(* Logix 5000 project; controller FV vendor 1 type 14 code 217 rev 31.11; software revision 31.00; part 24 of 63 *)
(* tags used below, declared in another part *)
   CheckTimeMask : INT;
   Delphi_Does_Eng_Func : BOOL;
   FR_FV30_AV01 : PlantItem;   // FV30_AV01
   FR_FV30_AV04 : PlantItem;   // FV30_AV04
   FR_FV30_AV05 : PlantItem;   // FV30_AV05
   FR_FV30_AV06 : PlantItem;   // FV30_AV06
   FR_FV30_AV07 : PlantItem;   // FV30_AV07
   FR_FV31_AV01 : PlantItem;   // FV31_AV01
   FR_N255 : INT[265];   // CHECKWORDS
   FR_VB4_AV17 : PlantItem;   // VB4_AV17
   FR_VB4_AV18 : PlantItem;   // VB4_AV18
   FR_VB4_AV19 : PlantItem;   // VB4_AV19
   FR_VB4_AV20 : PlantItem;   // VB4_AV20
   FR_VB4_AV21 : PlantItem;   // VB4_AV21
   FR_VB4_AV22 : PlantItem;   // VB4_AV22
   FR_VB4_AV23 : PlantItem;   // VB4_AV23
   TempChecktime : DINT;
(* FR_Common, continued *)

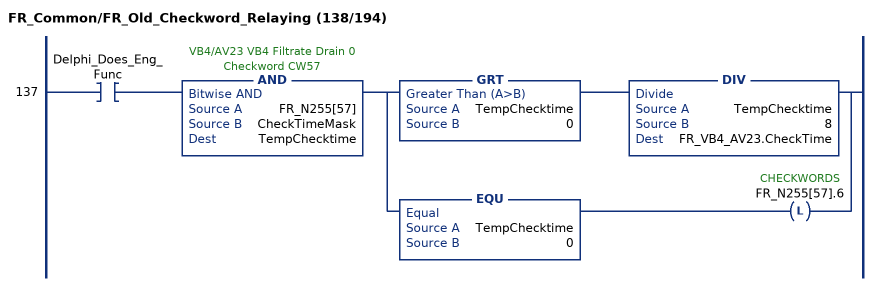
   [picture p442: FR_Common/FR_Old_Checkword_Relaying rungs 137-137]
   137: XIC(Delphi_Does_Eng_Func)AND(FR_N255[57],CheckTimeMask,TempChecktime)[GRT(TempChecktime,0) DIV(TempChecktime,8,FR_VB4_AV23.CheckTime) ,EQU(TempChecktime,0) OTL(FR_N255[57].6) ];
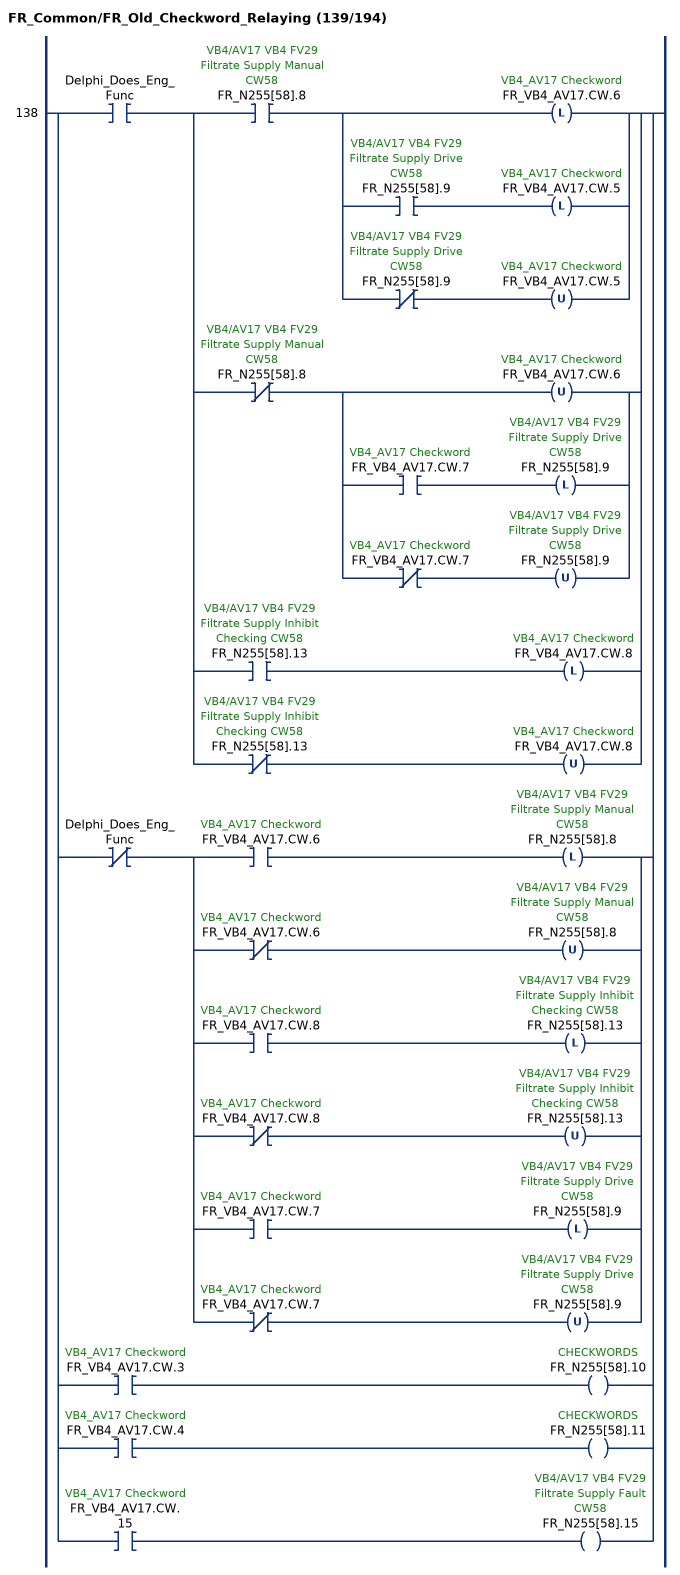
   138: [XIC(Delphi_Does_Eng_Func) [[XIC(FR_N255[58].8) [OTL(FR_VB4_AV17.CW.6) ,XIC(FR_N255[58].9) OTL(FR_VB4_AV17.CW.5) ,XIO(FR_N255[58].9) OTU(FR_VB4_AV17.CW.5) ] ,XIO(FR_N255[58].8) [OTU(FR_VB4_AV17.CW.6) ,[XIC(FR_VB4_AV17.CW.7) OTL(FR_N255[58].9) ,XIO(FR_VB4_AV17.CW.7) OTU(FR_N255[58].9) ] ] ] ,[XIC(FR_N255[58].13) OTL(FR_VB4_AV17.CW.8) ,XIO(FR_N255[58].13) OTU(FR_VB4_AV17.CW.8) ] ] ,XIO(Delphi_Does_Eng_Func) [[XIC(FR_VB4_AV17.CW.6) OTL(FR_N255[58].8) ,XIO(FR_VB4_AV17.CW.6) OTU(FR_N255[58].8) ] ,[XIC(FR_VB4_AV17.CW.8) OTL(FR_N255[58].13) ,XIO(FR_VB4_AV17.CW.8) OTU(FR_N255[58].13) ] ,[XIC(FR_VB4_AV17.CW.7) OTL(FR_N255[58].9) ,XIO(FR_VB4_AV17.CW.7) OTU(FR_N255[58].9) ] ] ,XIC(FR_VB4_AV17.CW.3) OTE(FR_N255[58].10) ,XIC(FR_VB4_AV17.CW.4) OTE(FR_N255[58].11) ,XIC(FR_VB4_AV17.CW.15) OTE(FR_N255[58].15) ];
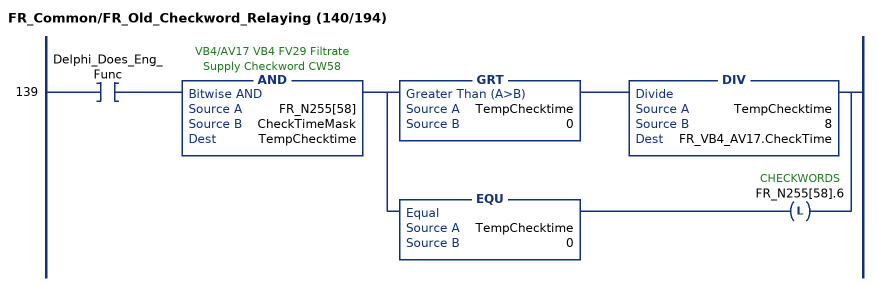
   139: XIC(Delphi_Does_Eng_Func)AND(FR_N255[58],CheckTimeMask,TempChecktime)[GRT(TempChecktime,0) DIV(TempChecktime,8,FR_VB4_AV17.CheckTime) ,EQU(TempChecktime,0) OTL(FR_N255[58].6) ];
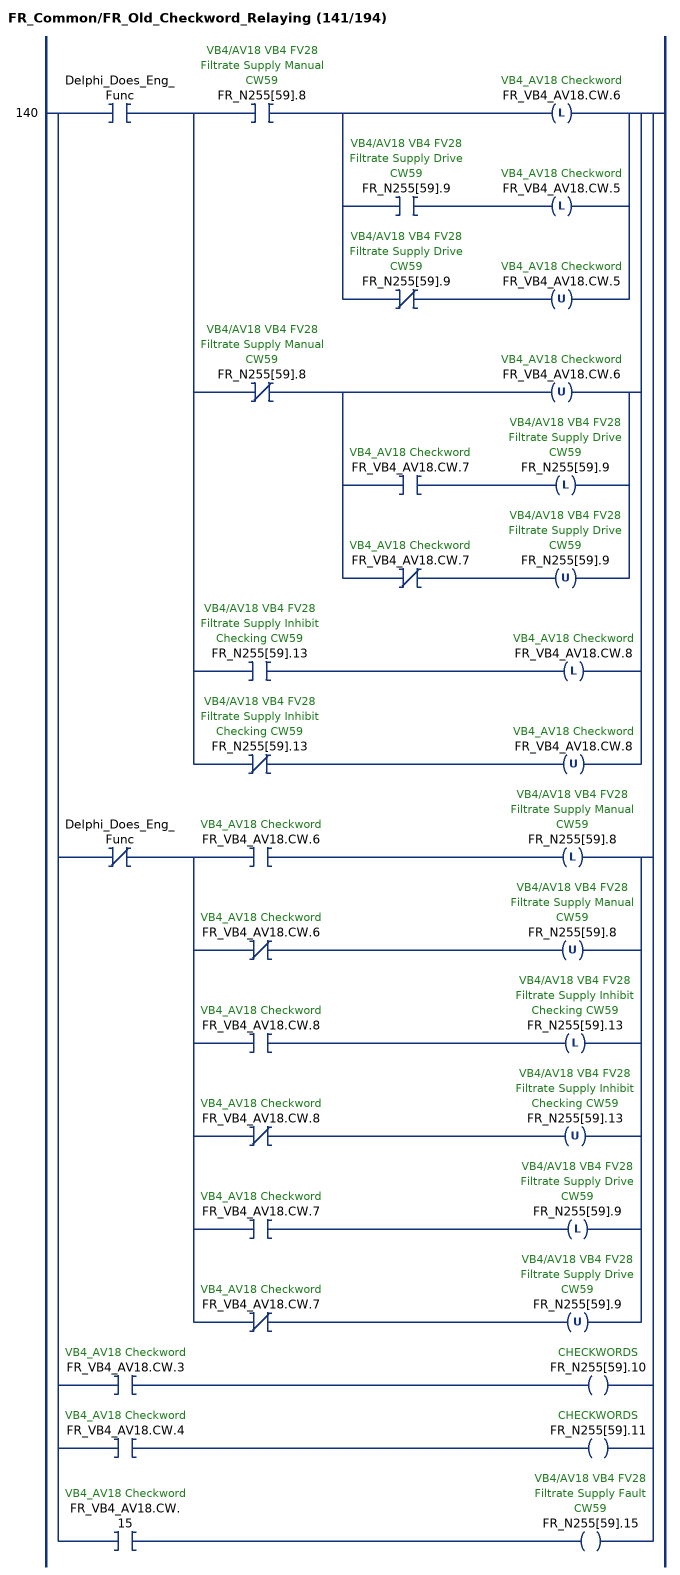
   140: [XIC(Delphi_Does_Eng_Func) [[XIC(FR_N255[59].8) [OTL(FR_VB4_AV18.CW.6) ,XIC(FR_N255[59].9) OTL(FR_VB4_AV18.CW.5) ,XIO(FR_N255[59].9) OTU(FR_VB4_AV18.CW.5) ] ,XIO(FR_N255[59].8) [OTU(FR_VB4_AV18.CW.6) ,[XIC(FR_VB4_AV18.CW.7) OTL(FR_N255[59].9) ,XIO(FR_VB4_AV18.CW.7) OTU(FR_N255[59].9) ] ] ] ,[XIC(FR_N255[59].13) OTL(FR_VB4_AV18.CW.8) ,XIO(FR_N255[59].13) OTU(FR_VB4_AV18.CW.8) ] ] ,XIO(Delphi_Does_Eng_Func) [[XIC(FR_VB4_AV18.CW.6) OTL(FR_N255[59].8) ,XIO(FR_VB4_AV18.CW.6) OTU(FR_N255[59].8) ] ,[XIC(FR_VB4_AV18.CW.8) OTL(FR_N255[59].13) ,XIO(FR_VB4_AV18.CW.8) OTU(FR_N255[59].13) ] ,[XIC(FR_VB4_AV18.CW.7) OTL(FR_N255[59].9) ,XIO(FR_VB4_AV18.CW.7) OTU(FR_N255[59].9) ] ] ,XIC(FR_VB4_AV18.CW.3) OTE(FR_N255[59].10) ,XIC(FR_VB4_AV18.CW.4) OTE(FR_N255[59].11) ,XIC(FR_VB4_AV18.CW.15) OTE(FR_N255[59].15) ];
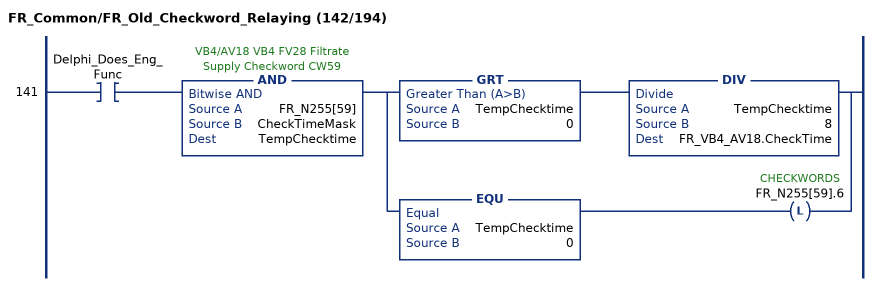
   141: XIC(Delphi_Does_Eng_Func)AND(FR_N255[59],CheckTimeMask,TempChecktime)[GRT(TempChecktime,0) DIV(TempChecktime,8,FR_VB4_AV18.CheckTime) ,EQU(TempChecktime,0) OTL(FR_N255[59].6) ];
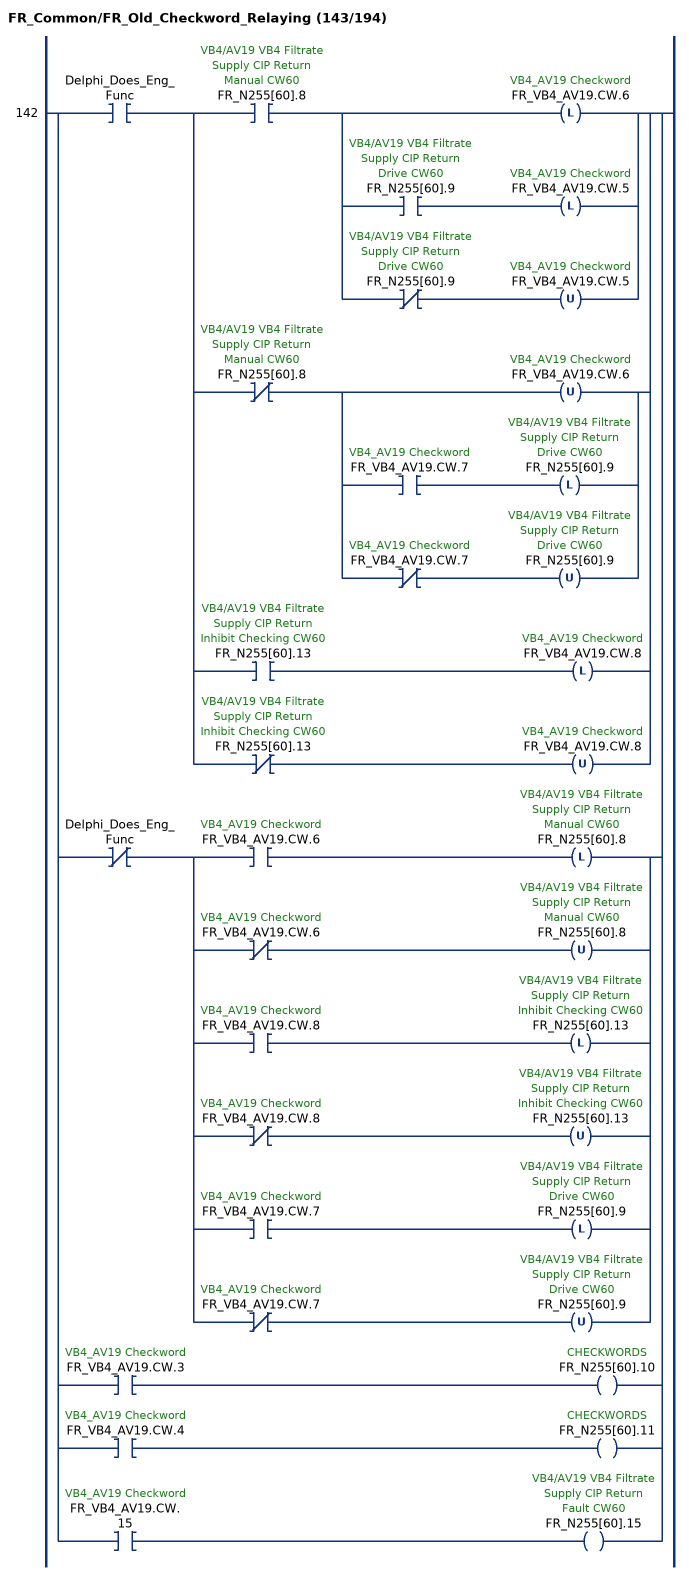
   142: [XIC(Delphi_Does_Eng_Func) [[XIC(FR_N255[60].8) [OTL(FR_VB4_AV19.CW.6) ,XIC(FR_N255[60].9) OTL(FR_VB4_AV19.CW.5) ,XIO(FR_N255[60].9) OTU(FR_VB4_AV19.CW.5) ] ,XIO(FR_N255[60].8) [OTU(FR_VB4_AV19.CW.6) ,[XIC(FR_VB4_AV19.CW.7) OTL(FR_N255[60].9) ,XIO(FR_VB4_AV19.CW.7) OTU(FR_N255[60].9) ] ] ] ,[XIC(FR_N255[60].13) OTL(FR_VB4_AV19.CW.8) ,XIO(FR_N255[60].13) OTU(FR_VB4_AV19.CW.8) ] ] ,XIO(Delphi_Does_Eng_Func) [[XIC(FR_VB4_AV19.CW.6) OTL(FR_N255[60].8) ,XIO(FR_VB4_AV19.CW.6) OTU(FR_N255[60].8) ] ,[XIC(FR_VB4_AV19.CW.8) OTL(FR_N255[60].13) ,XIO(FR_VB4_AV19.CW.8) OTU(FR_N255[60].13) ] ,[XIC(FR_VB4_AV19.CW.7) OTL(FR_N255[60].9) ,XIO(FR_VB4_AV19.CW.7) OTU(FR_N255[60].9) ] ] ,XIC(FR_VB4_AV19.CW.3) OTE(FR_N255[60].10) ,XIC(FR_VB4_AV19.CW.4) OTE(FR_N255[60].11) ,XIC(FR_VB4_AV19.CW.15) OTE(FR_N255[60].15) ];
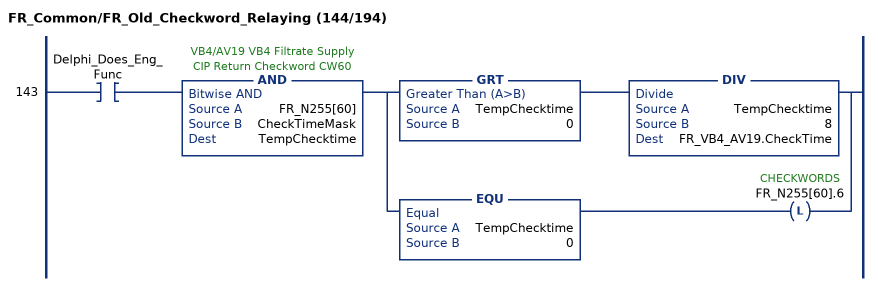
   143: XIC(Delphi_Does_Eng_Func)AND(FR_N255[60],CheckTimeMask,TempChecktime)[GRT(TempChecktime,0) DIV(TempChecktime,8,FR_VB4_AV19.CheckTime) ,EQU(TempChecktime,0) OTL(FR_N255[60].6) ];
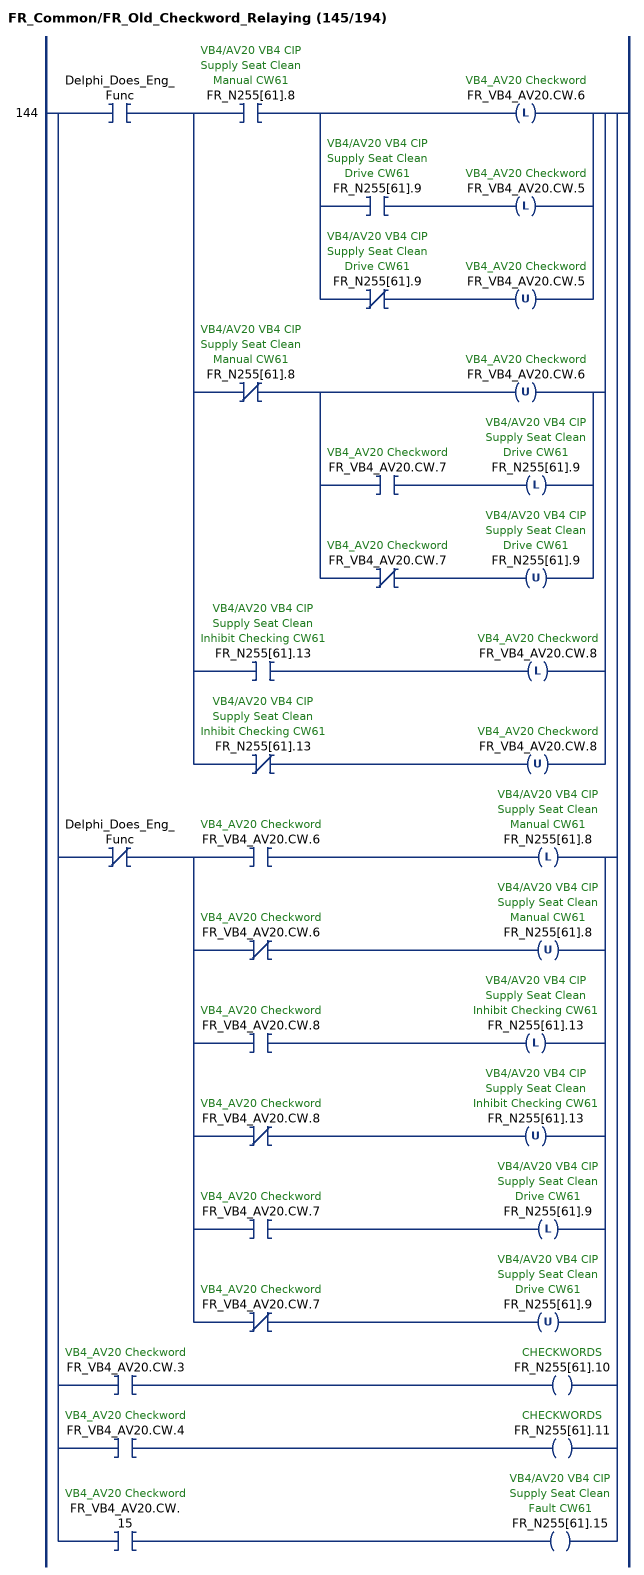
   144: [XIC(Delphi_Does_Eng_Func) [[XIC(FR_N255[61].8) [OTL(FR_VB4_AV20.CW.6) ,XIC(FR_N255[61].9) OTL(FR_VB4_AV20.CW.5) ,XIO(FR_N255[61].9) OTU(FR_VB4_AV20.CW.5) ] ,XIO(FR_N255[61].8) [OTU(FR_VB4_AV20.CW.6) ,[XIC(FR_VB4_AV20.CW.7) OTL(FR_N255[61].9) ,XIO(FR_VB4_AV20.CW.7) OTU(FR_N255[61].9) ] ] ] ,[XIC(FR_N255[61].13) OTL(FR_VB4_AV20.CW.8) ,XIO(FR_N255[61].13) OTU(FR_VB4_AV20.CW.8) ] ] ,XIO(Delphi_Does_Eng_Func) [[XIC(FR_VB4_AV20.CW.6) OTL(FR_N255[61].8) ,XIO(FR_VB4_AV20.CW.6) OTU(FR_N255[61].8) ] ,[XIC(FR_VB4_AV20.CW.8) OTL(FR_N255[61].13) ,XIO(FR_VB4_AV20.CW.8) OTU(FR_N255[61].13) ] ,[XIC(FR_VB4_AV20.CW.7) OTL(FR_N255[61].9) ,XIO(FR_VB4_AV20.CW.7) OTU(FR_N255[61].9) ] ] ,XIC(FR_VB4_AV20.CW.3) OTE(FR_N255[61].10) ,XIC(FR_VB4_AV20.CW.4) OTE(FR_N255[61].11) ,XIC(FR_VB4_AV20.CW.15) OTE(FR_N255[61].15) ];
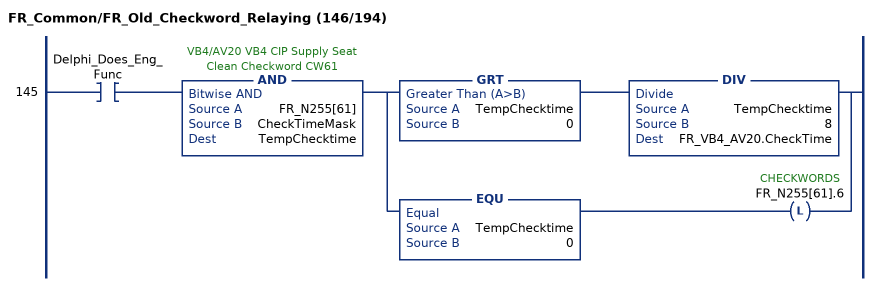
   145: XIC(Delphi_Does_Eng_Func)AND(FR_N255[61],CheckTimeMask,TempChecktime)[GRT(TempChecktime,0) DIV(TempChecktime,8,FR_VB4_AV20.CheckTime) ,EQU(TempChecktime,0) OTL(FR_N255[61].6) ];
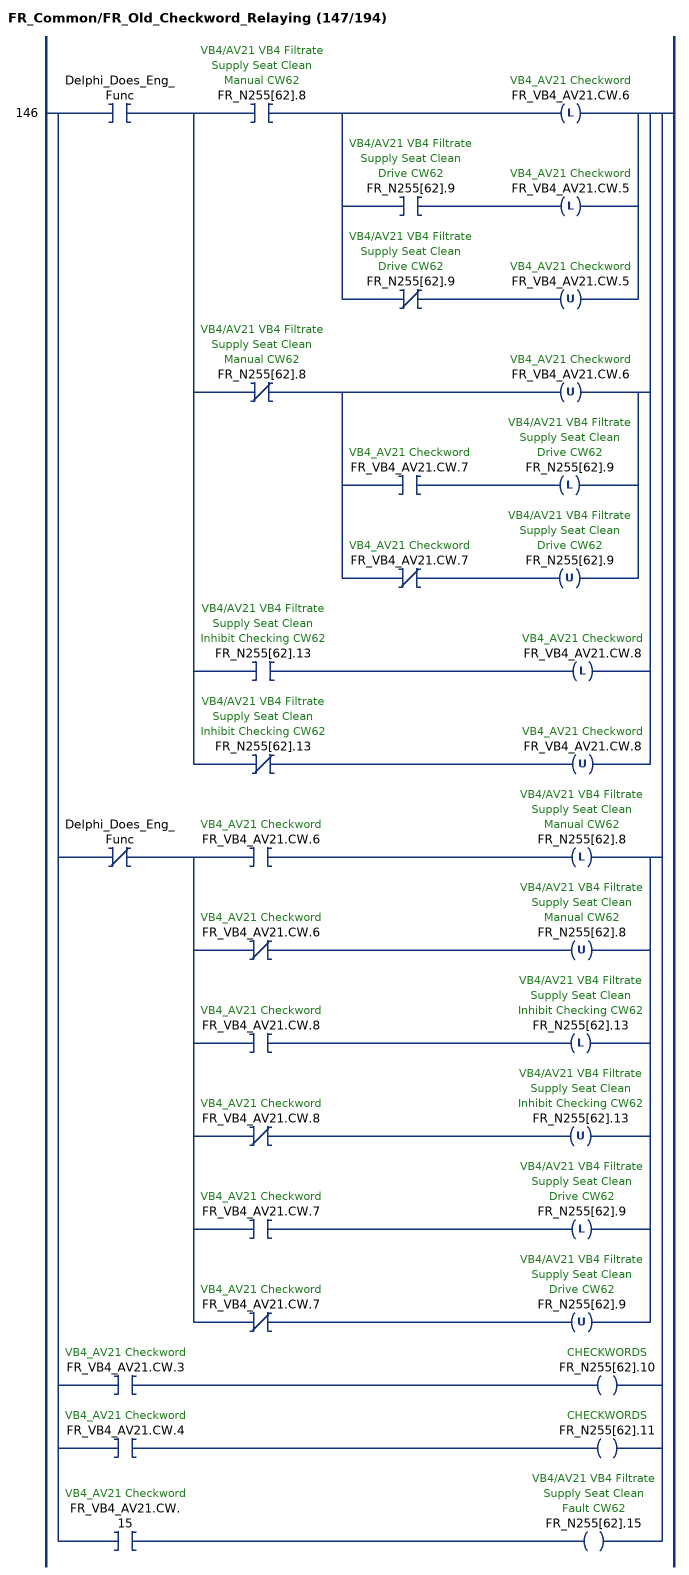
   146: [XIC(Delphi_Does_Eng_Func) [[XIC(FR_N255[62].8) [OTL(FR_VB4_AV21.CW.6) ,XIC(FR_N255[62].9) OTL(FR_VB4_AV21.CW.5) ,XIO(FR_N255[62].9) OTU(FR_VB4_AV21.CW.5) ] ,XIO(FR_N255[62].8) [OTU(FR_VB4_AV21.CW.6) ,[XIC(FR_VB4_AV21.CW.7) OTL(FR_N255[62].9) ,XIO(FR_VB4_AV21.CW.7) OTU(FR_N255[62].9) ] ] ] ,[XIC(FR_N255[62].13) OTL(FR_VB4_AV21.CW.8) ,XIO(FR_N255[62].13) OTU(FR_VB4_AV21.CW.8) ] ] ,XIO(Delphi_Does_Eng_Func) [[XIC(FR_VB4_AV21.CW.6) OTL(FR_N255[62].8) ,XIO(FR_VB4_AV21.CW.6) OTU(FR_N255[62].8) ] ,[XIC(FR_VB4_AV21.CW.8) OTL(FR_N255[62].13) ,XIO(FR_VB4_AV21.CW.8) OTU(FR_N255[62].13) ] ,[XIC(FR_VB4_AV21.CW.7) OTL(FR_N255[62].9) ,XIO(FR_VB4_AV21.CW.7) OTU(FR_N255[62].9) ] ] ,XIC(FR_VB4_AV21.CW.3) OTE(FR_N255[62].10) ,XIC(FR_VB4_AV21.CW.4) OTE(FR_N255[62].11) ,XIC(FR_VB4_AV21.CW.15) OTE(FR_N255[62].15) ];
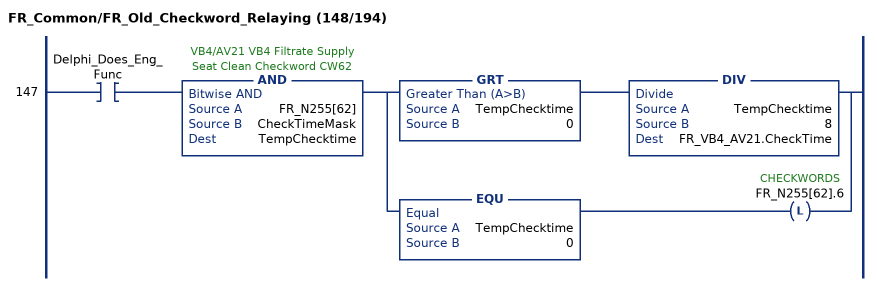
   147: XIC(Delphi_Does_Eng_Func)AND(FR_N255[62],CheckTimeMask,TempChecktime)[GRT(TempChecktime,0) DIV(TempChecktime,8,FR_VB4_AV21.CheckTime) ,EQU(TempChecktime,0) OTL(FR_N255[62].6) ];
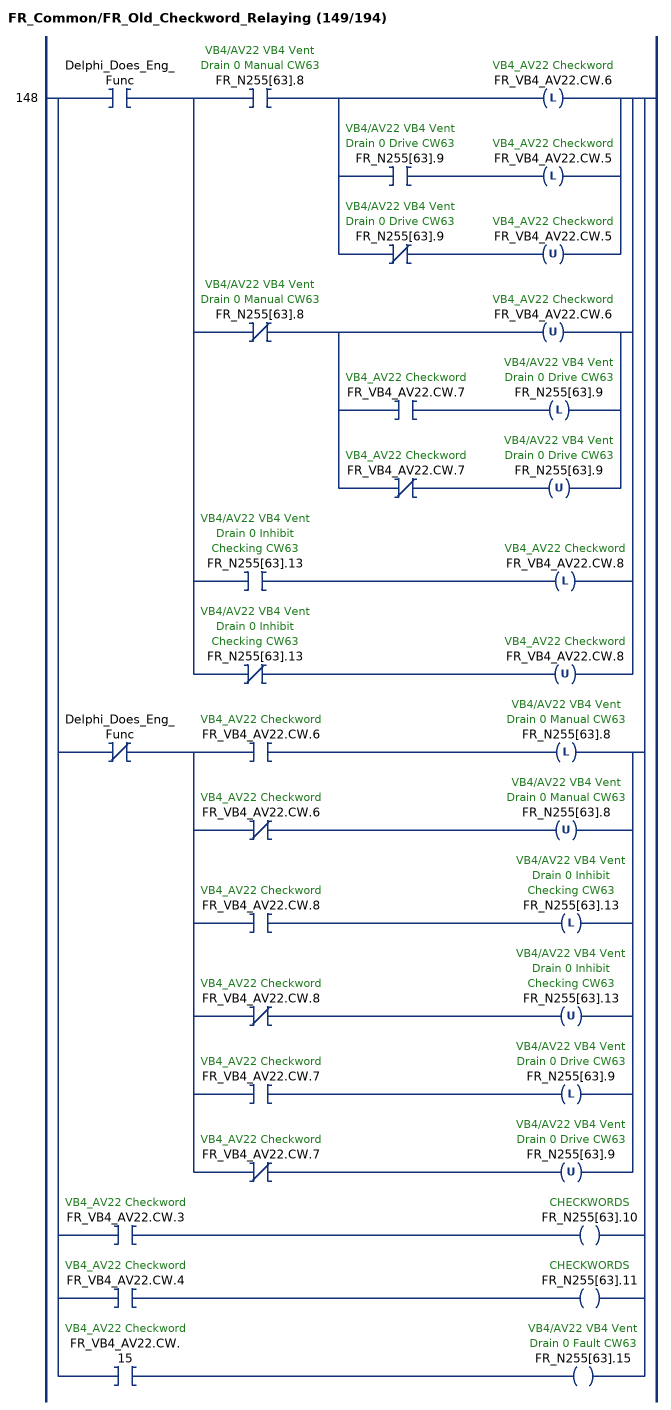
   148: [XIC(Delphi_Does_Eng_Func) [[XIC(FR_N255[63].8) [OTL(FR_VB4_AV22.CW.6) ,XIC(FR_N255[63].9) OTL(FR_VB4_AV22.CW.5) ,XIO(FR_N255[63].9) OTU(FR_VB4_AV22.CW.5) ] ,XIO(FR_N255[63].8) [OTU(FR_VB4_AV22.CW.6) ,[XIC(FR_VB4_AV22.CW.7) OTL(FR_N255[63].9) ,XIO(FR_VB4_AV22.CW.7) OTU(FR_N255[63].9) ] ] ] ,[XIC(FR_N255[63].13) OTL(FR_VB4_AV22.CW.8) ,XIO(FR_N255[63].13) OTU(FR_VB4_AV22.CW.8) ] ] ,XIO(Delphi_Does_Eng_Func) [[XIC(FR_VB4_AV22.CW.6) OTL(FR_N255[63].8) ,XIO(FR_VB4_AV22.CW.6) OTU(FR_N255[63].8) ] ,[XIC(FR_VB4_AV22.CW.8) OTL(FR_N255[63].13) ,XIO(FR_VB4_AV22.CW.8) OTU(FR_N255[63].13) ] ,[XIC(FR_VB4_AV22.CW.7) OTL(FR_N255[63].9) ,XIO(FR_VB4_AV22.CW.7) OTU(FR_N255[63].9) ] ] ,XIC(FR_VB4_AV22.CW.3) OTE(FR_N255[63].10) ,XIC(FR_VB4_AV22.CW.4) OTE(FR_N255[63].11) ,XIC(FR_VB4_AV22.CW.15) OTE(FR_N255[63].15) ];
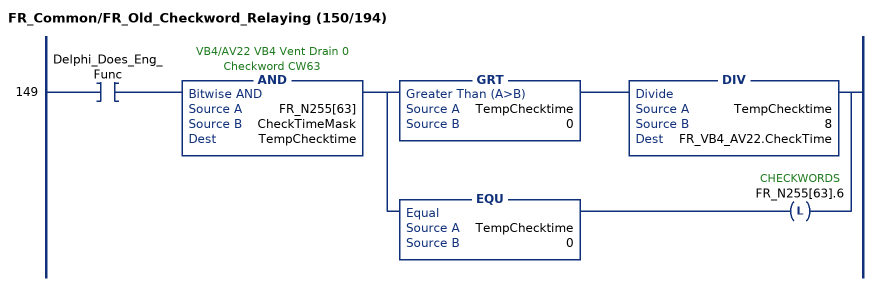
   149: XIC(Delphi_Does_Eng_Func)AND(FR_N255[63],CheckTimeMask,TempChecktime)[GRT(TempChecktime,0) DIV(TempChecktime,8,FR_VB4_AV22.CheckTime) ,EQU(TempChecktime,0) OTL(FR_N255[63].6) ];
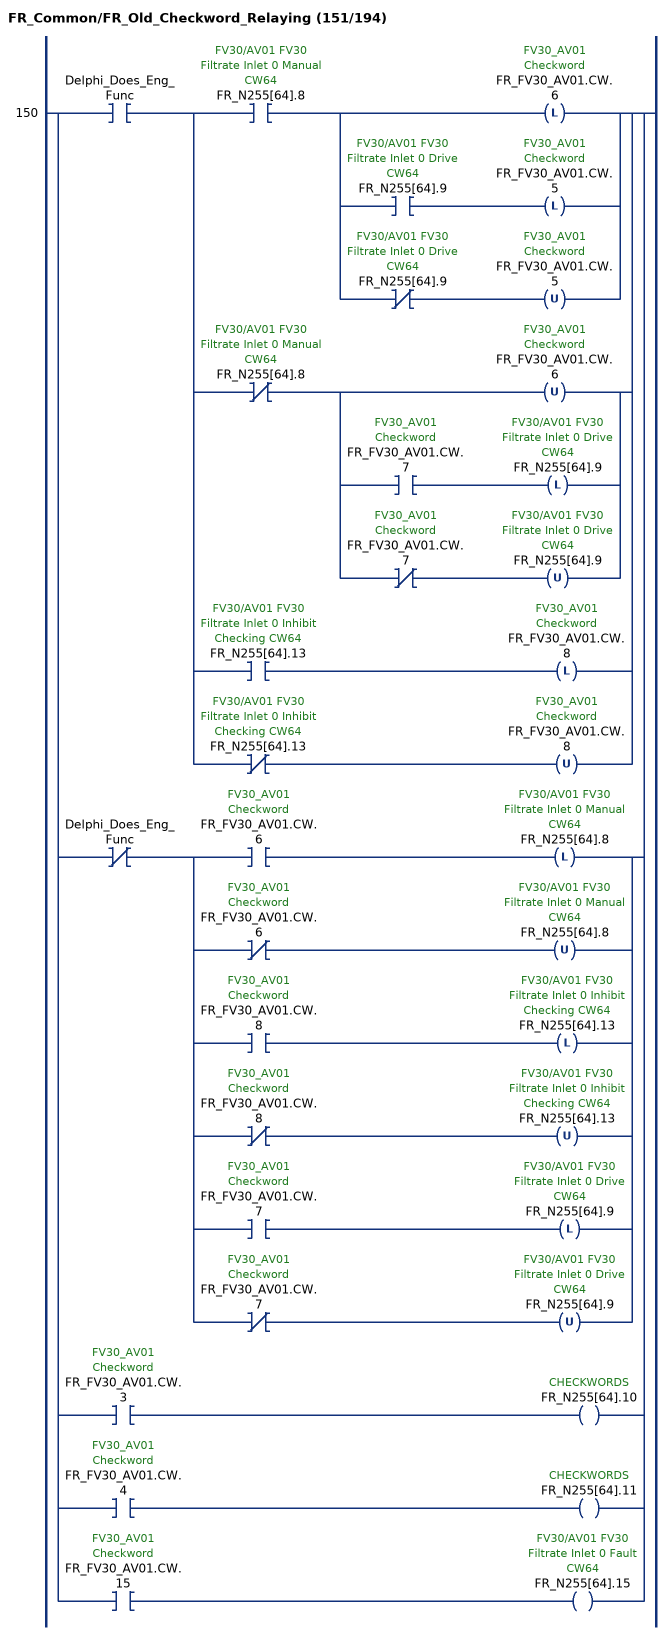
   150: [XIC(Delphi_Does_Eng_Func) [[XIC(FR_N255[64].8) [OTL(FR_FV30_AV01.CW.6) ,XIC(FR_N255[64].9) OTL(FR_FV30_AV01.CW.5) ,XIO(FR_N255[64].9) OTU(FR_FV30_AV01.CW.5) ] ,XIO(FR_N255[64].8) [OTU(FR_FV30_AV01.CW.6) ,[XIC(FR_FV30_AV01.CW.7) OTL(FR_N255[64].9) ,XIO(FR_FV30_AV01.CW.7) OTU(FR_N255[64].9) ] ] ] ,[XIC(FR_N255[64].13) OTL(FR_FV30_AV01.CW.8) ,XIO(FR_N255[64].13) OTU(FR_FV30_AV01.CW.8) ] ] ,XIO(Delphi_Does_Eng_Func) [[XIC(FR_FV30_AV01.CW.6) OTL(FR_N255[64].8) ,XIO(FR_FV30_AV01.CW.6) OTU(FR_N255[64].8) ] ,[XIC(FR_FV30_AV01.CW.8) OTL(FR_N255[64].13) ,XIO(FR_FV30_AV01.CW.8) OTU(FR_N255[64].13) ] ,[XIC(FR_FV30_AV01.CW.7) OTL(FR_N255[64].9) ,XIO(FR_FV30_AV01.CW.7) OTU(FR_N255[64].9) ] ] ,XIC(FR_FV30_AV01.CW.3) OTE(FR_N255[64].10) ,XIC(FR_FV30_AV01.CW.4) OTE(FR_N255[64].11) ,XIC(FR_FV30_AV01.CW.15) OTE(FR_N255[64].15) ];
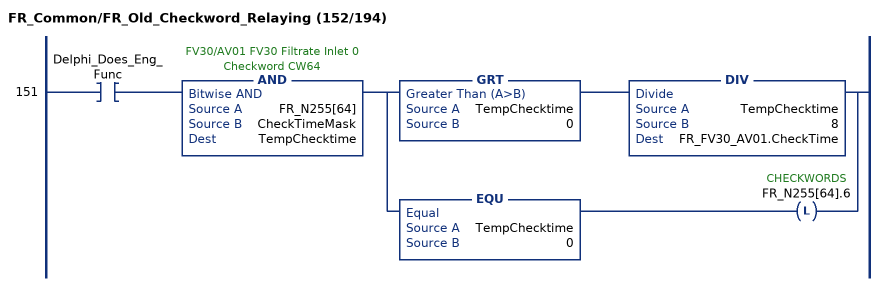
   151: XIC(Delphi_Does_Eng_Func)AND(FR_N255[64],CheckTimeMask,TempChecktime)[GRT(TempChecktime,0) DIV(TempChecktime,8,FR_FV30_AV01.CheckTime) ,EQU(TempChecktime,0) OTL(FR_N255[64].6) ];
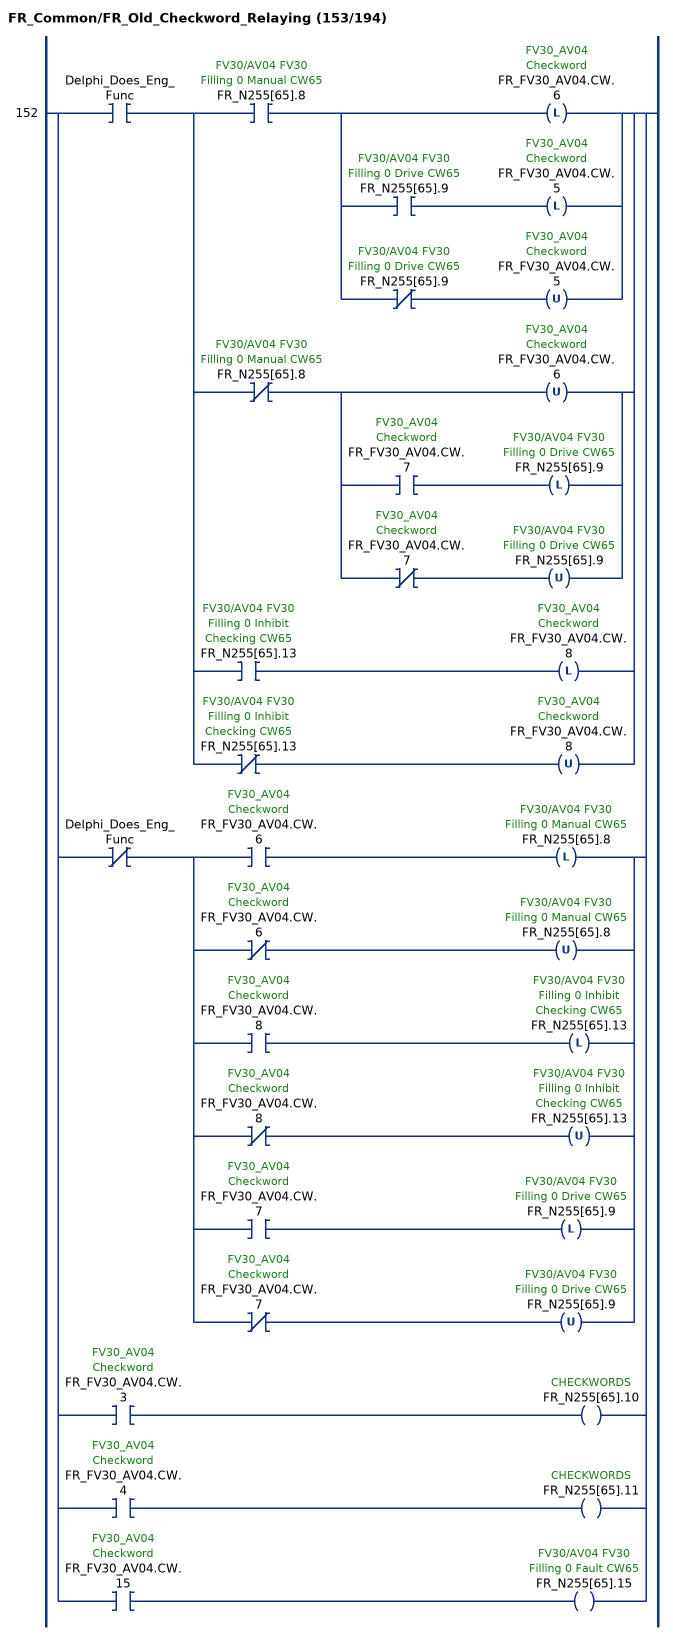
   152: [XIC(Delphi_Does_Eng_Func) [[XIC(FR_N255[65].8) [OTL(FR_FV30_AV04.CW.6) ,XIC(FR_N255[65].9) OTL(FR_FV30_AV04.CW.5) ,XIO(FR_N255[65].9) OTU(FR_FV30_AV04.CW.5) ] ,XIO(FR_N255[65].8) [OTU(FR_FV30_AV04.CW.6) ,[XIC(FR_FV30_AV04.CW.7) OTL(FR_N255[65].9) ,XIO(FR_FV30_AV04.CW.7) OTU(FR_N255[65].9) ] ] ] ,[XIC(FR_N255[65].13) OTL(FR_FV30_AV04.CW.8) ,XIO(FR_N255[65].13) OTU(FR_FV30_AV04.CW.8) ] ] ,XIO(Delphi_Does_Eng_Func) [[XIC(FR_FV30_AV04.CW.6) OTL(FR_N255[65].8) ,XIO(FR_FV30_AV04.CW.6) OTU(FR_N255[65].8) ] ,[XIC(FR_FV30_AV04.CW.8) OTL(FR_N255[65].13) ,XIO(FR_FV30_AV04.CW.8) OTU(FR_N255[65].13) ] ,[XIC(FR_FV30_AV04.CW.7) OTL(FR_N255[65].9) ,XIO(FR_FV30_AV04.CW.7) OTU(FR_N255[65].9) ] ] ,XIC(FR_FV30_AV04.CW.3) OTE(FR_N255[65].10) ,XIC(FR_FV30_AV04.CW.4) OTE(FR_N255[65].11) ,XIC(FR_FV30_AV04.CW.15) OTE(FR_N255[65].15) ];
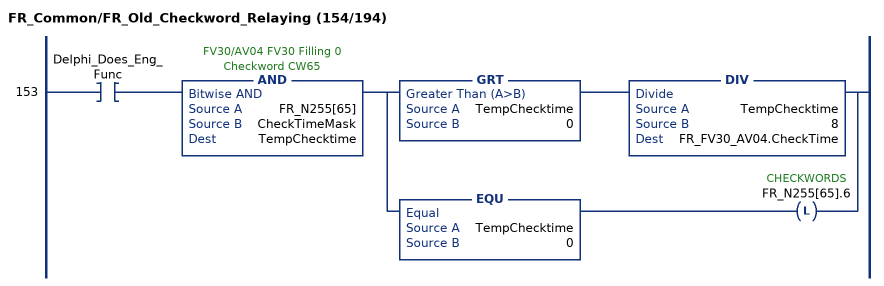
   153: XIC(Delphi_Does_Eng_Func)AND(FR_N255[65],CheckTimeMask,TempChecktime)[GRT(TempChecktime,0) DIV(TempChecktime,8,FR_FV30_AV04.CheckTime) ,EQU(TempChecktime,0) OTL(FR_N255[65].6) ];
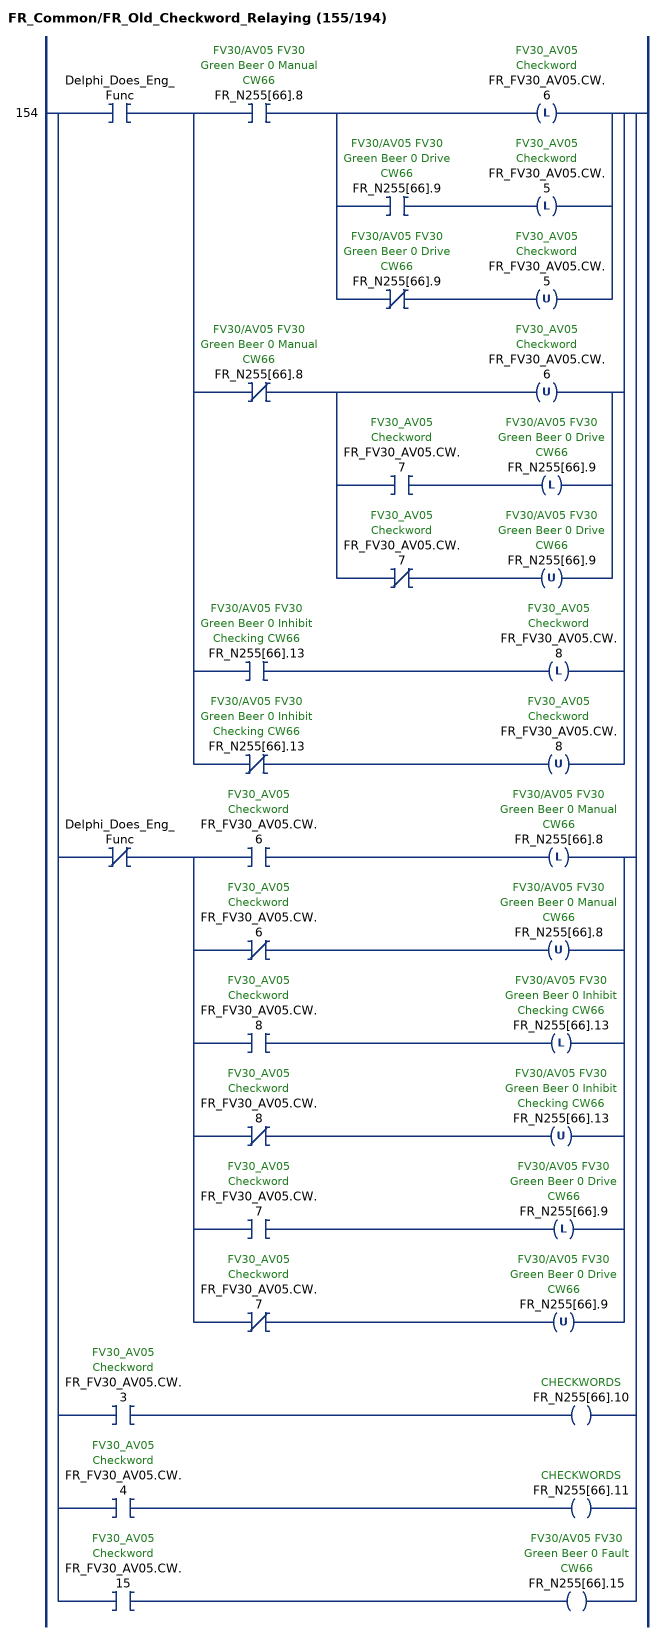
   154: [XIC(Delphi_Does_Eng_Func) [[XIC(FR_N255[66].8) [OTL(FR_FV30_AV05.CW.6) ,XIC(FR_N255[66].9) OTL(FR_FV30_AV05.CW.5) ,XIO(FR_N255[66].9) OTU(FR_FV30_AV05.CW.5) ] ,XIO(FR_N255[66].8) [OTU(FR_FV30_AV05.CW.6) ,[XIC(FR_FV30_AV05.CW.7) OTL(FR_N255[66].9) ,XIO(FR_FV30_AV05.CW.7) OTU(FR_N255[66].9) ] ] ] ,[XIC(FR_N255[66].13) OTL(FR_FV30_AV05.CW.8) ,XIO(FR_N255[66].13) OTU(FR_FV30_AV05.CW.8) ] ] ,XIO(Delphi_Does_Eng_Func) [[XIC(FR_FV30_AV05.CW.6) OTL(FR_N255[66].8) ,XIO(FR_FV30_AV05.CW.6) OTU(FR_N255[66].8) ] ,[XIC(FR_FV30_AV05.CW.8) OTL(FR_N255[66].13) ,XIO(FR_FV30_AV05.CW.8) OTU(FR_N255[66].13) ] ,[XIC(FR_FV30_AV05.CW.7) OTL(FR_N255[66].9) ,XIO(FR_FV30_AV05.CW.7) OTU(FR_N255[66].9) ] ] ,XIC(FR_FV30_AV05.CW.3) OTE(FR_N255[66].10) ,XIC(FR_FV30_AV05.CW.4) OTE(FR_N255[66].11) ,XIC(FR_FV30_AV05.CW.15) OTE(FR_N255[66].15) ];
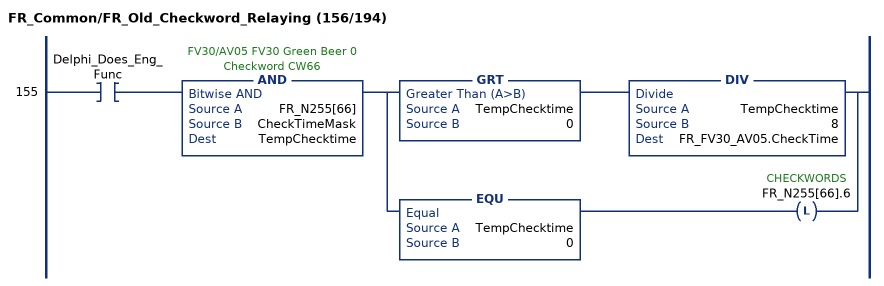
   155: XIC(Delphi_Does_Eng_Func)AND(FR_N255[66],CheckTimeMask,TempChecktime)[GRT(TempChecktime,0) DIV(TempChecktime,8,FR_FV30_AV05.CheckTime) ,EQU(TempChecktime,0) OTL(FR_N255[66].6) ];
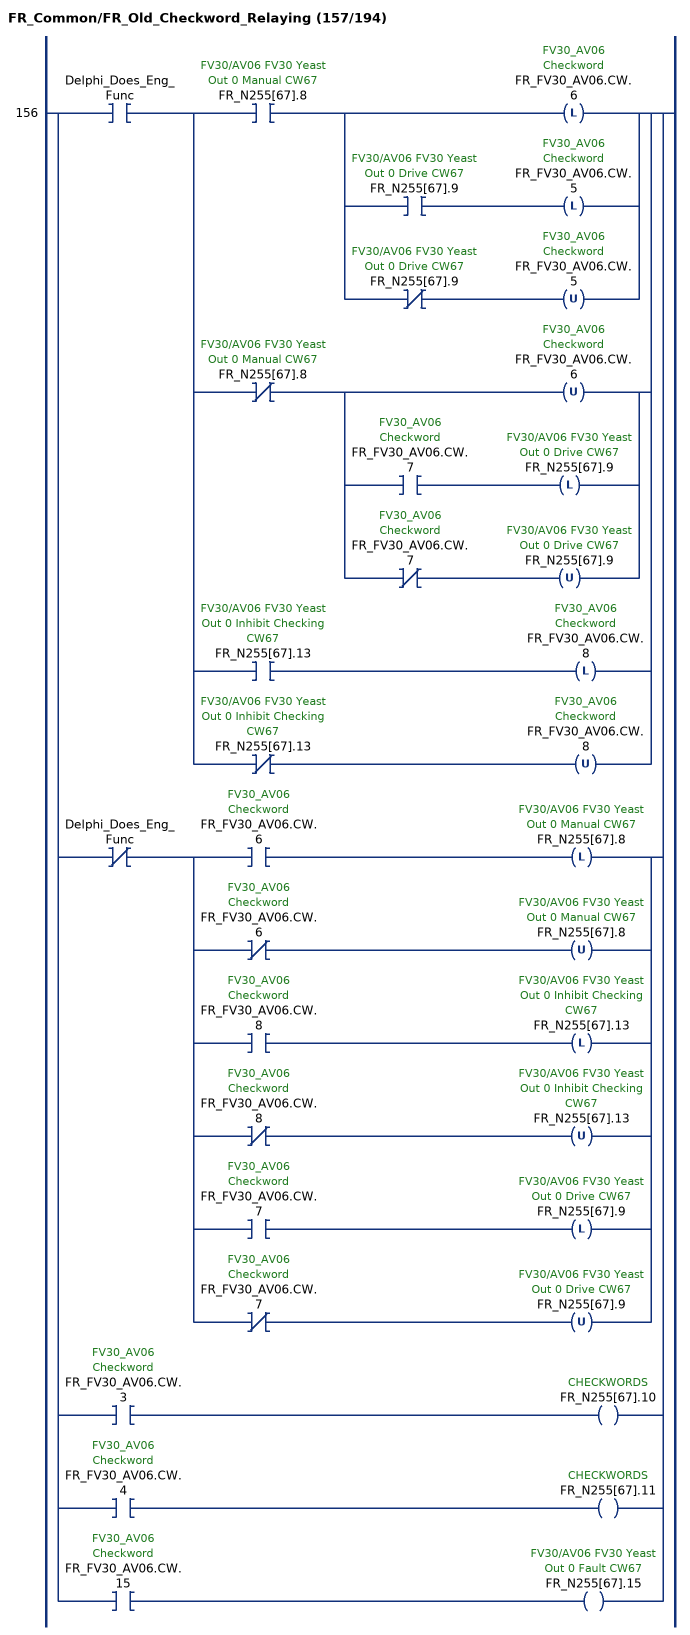
   156: [XIC(Delphi_Does_Eng_Func) [[XIC(FR_N255[67].8) [OTL(FR_FV30_AV06.CW.6) ,XIC(FR_N255[67].9) OTL(FR_FV30_AV06.CW.5) ,XIO(FR_N255[67].9) OTU(FR_FV30_AV06.CW.5) ] ,XIO(FR_N255[67].8) [OTU(FR_FV30_AV06.CW.6) ,[XIC(FR_FV30_AV06.CW.7) OTL(FR_N255[67].9) ,XIO(FR_FV30_AV06.CW.7) OTU(FR_N255[67].9) ] ] ] ,[XIC(FR_N255[67].13) OTL(FR_FV30_AV06.CW.8) ,XIO(FR_N255[67].13) OTU(FR_FV30_AV06.CW.8) ] ] ,XIO(Delphi_Does_Eng_Func) [[XIC(FR_FV30_AV06.CW.6) OTL(FR_N255[67].8) ,XIO(FR_FV30_AV06.CW.6) OTU(FR_N255[67].8) ] ,[XIC(FR_FV30_AV06.CW.8) OTL(FR_N255[67].13) ,XIO(FR_FV30_AV06.CW.8) OTU(FR_N255[67].13) ] ,[XIC(FR_FV30_AV06.CW.7) OTL(FR_N255[67].9) ,XIO(FR_FV30_AV06.CW.7) OTU(FR_N255[67].9) ] ] ,XIC(FR_FV30_AV06.CW.3) OTE(FR_N255[67].10) ,XIC(FR_FV30_AV06.CW.4) OTE(FR_N255[67].11) ,XIC(FR_FV30_AV06.CW.15) OTE(FR_N255[67].15) ];
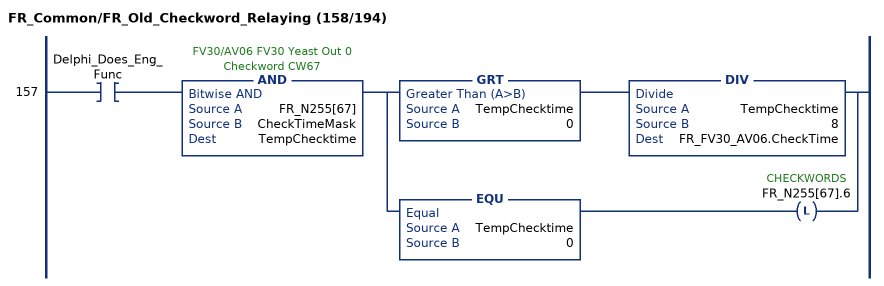
   157: XIC(Delphi_Does_Eng_Func)AND(FR_N255[67],CheckTimeMask,TempChecktime)[GRT(TempChecktime,0) DIV(TempChecktime,8,FR_FV30_AV06.CheckTime) ,EQU(TempChecktime,0) OTL(FR_N255[67].6) ];
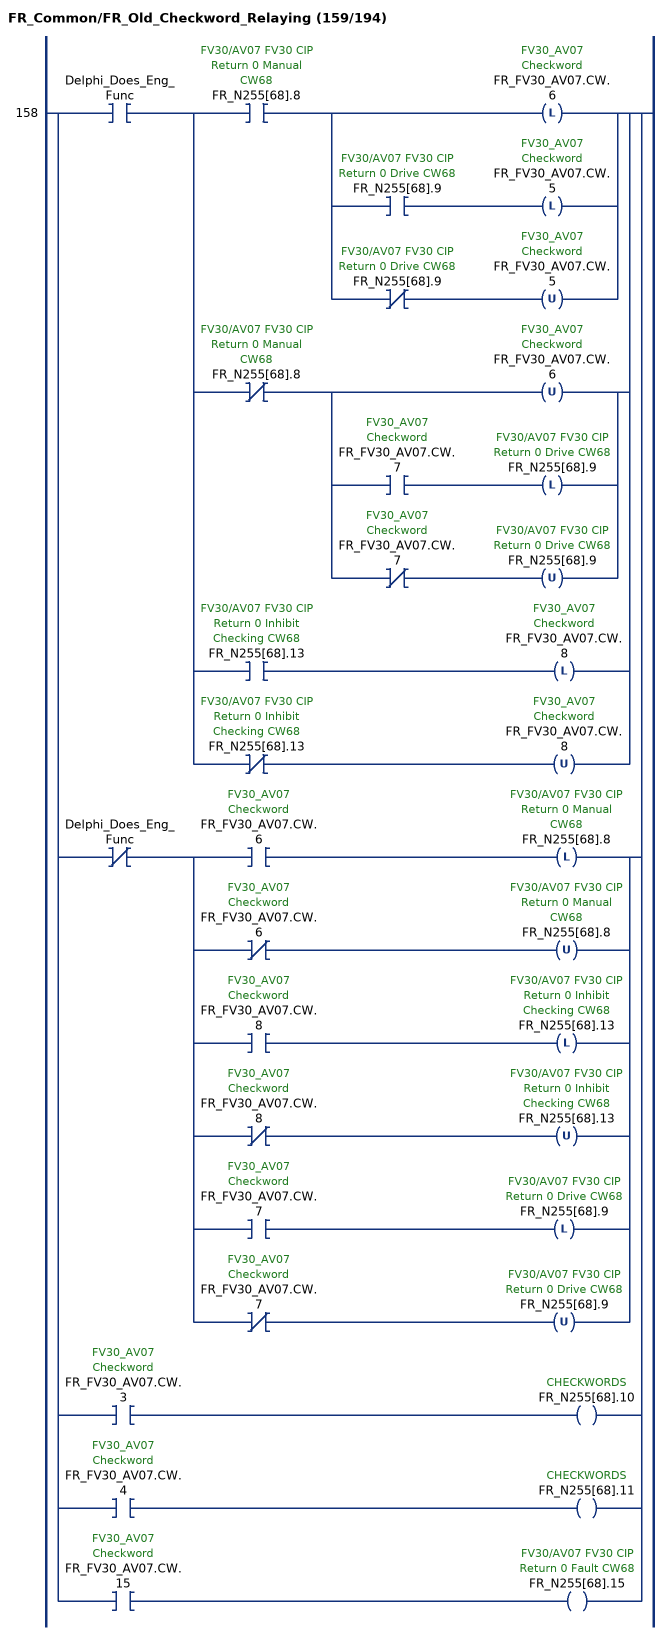
   158: [XIC(Delphi_Does_Eng_Func) [[XIC(FR_N255[68].8) [OTL(FR_FV30_AV07.CW.6) ,XIC(FR_N255[68].9) OTL(FR_FV30_AV07.CW.5) ,XIO(FR_N255[68].9) OTU(FR_FV30_AV07.CW.5) ] ,XIO(FR_N255[68].8) [OTU(FR_FV30_AV07.CW.6) ,[XIC(FR_FV30_AV07.CW.7) OTL(FR_N255[68].9) ,XIO(FR_FV30_AV07.CW.7) OTU(FR_N255[68].9) ] ] ] ,[XIC(FR_N255[68].13) OTL(FR_FV30_AV07.CW.8) ,XIO(FR_N255[68].13) OTU(FR_FV30_AV07.CW.8) ] ] ,XIO(Delphi_Does_Eng_Func) [[XIC(FR_FV30_AV07.CW.6) OTL(FR_N255[68].8) ,XIO(FR_FV30_AV07.CW.6) OTU(FR_N255[68].8) ] ,[XIC(FR_FV30_AV07.CW.8) OTL(FR_N255[68].13) ,XIO(FR_FV30_AV07.CW.8) OTU(FR_N255[68].13) ] ,[XIC(FR_FV30_AV07.CW.7) OTL(FR_N255[68].9) ,XIO(FR_FV30_AV07.CW.7) OTU(FR_N255[68].9) ] ] ,XIC(FR_FV30_AV07.CW.3) OTE(FR_N255[68].10) ,XIC(FR_FV30_AV07.CW.4) OTE(FR_N255[68].11) ,XIC(FR_FV30_AV07.CW.15) OTE(FR_N255[68].15) ];
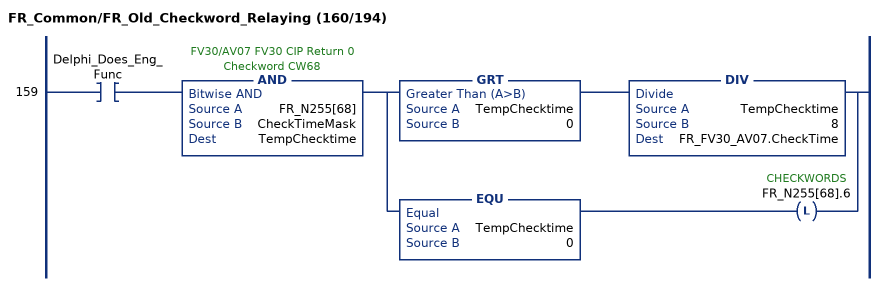
   159: XIC(Delphi_Does_Eng_Func)AND(FR_N255[68],CheckTimeMask,TempChecktime)[GRT(TempChecktime,0) DIV(TempChecktime,8,FR_FV30_AV07.CheckTime) ,EQU(TempChecktime,0) OTL(FR_N255[68].6) ];
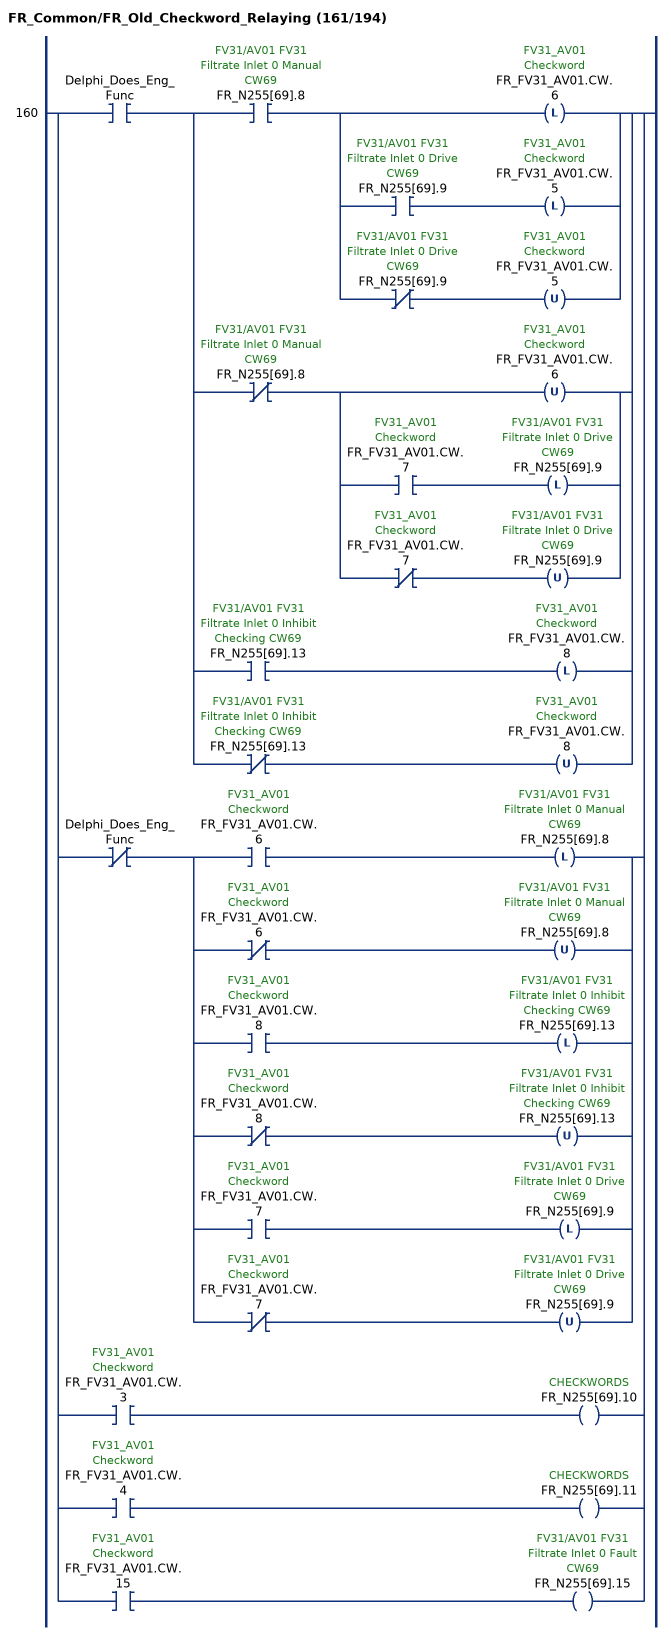
   160: [XIC(Delphi_Does_Eng_Func) [[XIC(FR_N255[69].8) [OTL(FR_FV31_AV01.CW.6) ,XIC(FR_N255[69].9) OTL(FR_FV31_AV01.CW.5) ,XIO(FR_N255[69].9) OTU(FR_FV31_AV01.CW.5) ] ,XIO(FR_N255[69].8) [OTU(FR_FV31_AV01.CW.6) ,[XIC(FR_FV31_AV01.CW.7) OTL(FR_N255[69].9) ,XIO(FR_FV31_AV01.CW.7) OTU(FR_N255[69].9) ] ] ] ,[XIC(FR_N255[69].13) OTL(FR_FV31_AV01.CW.8) ,XIO(FR_N255[69].13) OTU(FR_FV31_AV01.CW.8) ] ] ,XIO(Delphi_Does_Eng_Func) [[XIC(FR_FV31_AV01.CW.6) OTL(FR_N255[69].8) ,XIO(FR_FV31_AV01.CW.6) OTU(FR_N255[69].8) ] ,[XIC(FR_FV31_AV01.CW.8) OTL(FR_N255[69].13) ,XIO(FR_FV31_AV01.CW.8) OTU(FR_N255[69].13) ] ,[XIC(FR_FV31_AV01.CW.7) OTL(FR_N255[69].9) ,XIO(FR_FV31_AV01.CW.7) OTU(FR_N255[69].9) ] ] ,XIC(FR_FV31_AV01.CW.3) OTE(FR_N255[69].10) ,XIC(FR_FV31_AV01.CW.4) OTE(FR_N255[69].11) ,XIC(FR_FV31_AV01.CW.15) OTE(FR_N255[69].15) ];
